REGION Network 11: Habilita cambiar de CAPA_Elem_2
         OPN   "DB_Receta_Actual";
         SET;
         R     #Habil_2_CAPA;
         L     #Capa_Actual;
         L     #Max_Nro_Capas;
         >=I;
         JC    No2CAPA;
         L     #Adress_Capa;
         L     #Length_Capas;
         +I;
         L     #Offset_Filas_DB;
         +I;
         SLD   3;
         L     #Offset_Elementos_DB_bit;
         +I;
         L     #Length_Elementos_DB_bit;
         +I;
         LAR2;
         O     DBX [AR2, P#0.0];
         O     DBX [ AR2 , P#2.0 ];
         =     #Habil_2_CAPA;
   No2CAPA:NOP   0;
END_REGION

REGION Network 12: #Elemento_Actual
         OPN   "DB_Receta_Actual";

         A     DBX [ AR1 , P#4.0 ];
         =     #Elemento_Actual;

         A     #Elemento_Actual;
         JCN   NoActual;
         TAR1  AR2;
END_REGION

REGION Network 13: NUM = 1
         SET;
   // R DBX [ AR1 , P#4.0 ]
         A     #Habil_1_IZQ;
         JCN   No_1_IZQ;

         TAR1  AR2;
         L     1;
         +AR2;
   //S DBX [ AR2 , P#4.0 ]
         JU    Fin;

   No_1_IZQ:A     #Habil_1_ABA;
         JCN   No_ABA;
         L     #Adress_Filas_DB_bit;
         SRD   3;
         L     #Length_Filas_DB;
         +I;
         SLD   3;
         L     #Offset_Elementos_DB_bit;
         +I;
         LAR2;
         SET;
   //S DBX [ AR2 , P#4.0 ]
         JU    Fin;

   No_ABA:A     #Habil_1_CAPA;
         JCN   No_CAPA;
         L     #Adress_Capa;
         L     #Length_Capas;
         +I;
         L     #Offset_Filas_DB;
         +I;
         SLD   3;
         L     #Offset_Elementos_DB_bit;
         +I;
         LAR2;
   //S DBX [ AR2 , P#4.0 ]
         L     #Capa_Actual;
         L     1;
         +I;
         T     #Capa_Actual;
         JU    Fin;

   No_CAPA:NOP   0;
         L     #Offset_Capas;
         L     #Offset_Filas_DB;
         +I;
         SLD   3;
         L     #Offset_Elementos_DB_bit;
         +I;
         LAR2;
   //S DBX [ AR2 , P#4.0 ]
         L     1;
         T     #Capa_Actual;
         L     #Nro_Pallet;
         L     1;
         +I;
         T     #Nro_Pallet;
         JU    Fin;
END_REGION

REGION Network 14: No elemento actual
   NoNUM:JU    Fin;
   NoActual:NOP   0;
END_REGION

REGION Network 15: Bucle Elementos
         L     #Índice_Elementos;
         L     1;
         +I;
         T     #Índice_Elementos;
         L     #Max_Nro_Elementos;
         <=I;
         JC    New_Ele;
END_REGION

REGION Network 16: Bucle Filas
         L     1;
         T     #Índice_Elementos;
         L     #Índice_Filas;
         L     1;
         +I;
         T     #Índice_Filas;
         L     #Max_Nro_Filas;
         <=I;
         JC    New_Fil;
END_REGION

REGION Network 17: #Error
         SET;
         S     #Error;
END_REGION

REGION Network 18: Fin de Bloque
   Fin:  SET;
         R     #Error;
         OPN   "DB_Receta_Actual";
         AN    DBX [ AR2 , P#0.0 ];
         AN    DBX [ AR2 , P#2.0 ];
         JCN   NO_0;
         L     0;
         JU    Transferir;
   NO_0: A     DBX [ AR2 , P#0.0 ];
         AN    DBX [ AR2 , P#2.0 ];
         JCN   NO_1;
         L     1;
         JU    Transferir;
   NO_1: AN    DBX [ AR2 , P#0.0 ];
         A     DBX [ AR2 , P#2.0 ];
         JCN   NO_2;
         L     2;
         JU    Transferir;
   NO_2: L     3;
   Transferir:T     "Proceso Dosificador".Elemento_Proximo;
   // 0 = Invisible
   // 1 = V
   // 2 = H
   // 3 = HH
END_REGION
END_FUNCTION

FUNCTION "FC_Animación" : Void   // FC3, STL
{ S7_Optimized_Access := 'FALSE' }
VERSION : 0.1
BEGIN

REGION Network 1
         O     "Cambio_Elemento";
         O     "flanco"."nHMI.Pls_Inc_Capa";
         O     "flanco"."nHMI.Pls_Dec_Capa";
         O     "flanco"."pHMI.Pls_Inc_Capa_Editando";
         O     "flanco"."pHMI.Pls_Dec_Capa_Editando";

         =     #Cambio_Elemento;
END_REGION

REGION Network 2: Inicializa fila y elemento
         A     "CicIni";
         JCN   L001;
         L     1;
         T     "DB_Animación".Elemento_SEL;
         T     "DB_Animación".Fila_SEL;
         L     "Puntero".Offset_Filas_HMI;
         L     "Puntero".Offset_Elementos_HMI;
         +I;
         SLD   3;
         LAR1;
         OPN   "DB_Animación";
         L     3;
         T     DBB [ AR1 , P#0.0 ];
         S     #Cambio_Elemento;
   L001: NOP   0;

         L     "DB_Animación".Fila_SEL;
         L     "DB_Animación".Elemento_SEL;
   // OFFSET_Y "0" en la primer fila
         L     "Puntero".Offset_Filas_HMI;
         OPN   "DB_Animación";
         SLD   3;
         LAR1;
         L     0;
         T     DBW [ AR1 , P#0.0 ];


   // OFFSET_X "0" en el primer elemento de la primer fila
         L     "Puntero".Offset_Filas_HMI;
         L     "Puntero".Offset_Elementos_HMI;
         +I;
         OPN   "DB_Animación";
         SLD   3;
         LAR1;
         L     0;
         T     DBW [ AR1 , P#2.0 ];

   //Edita recetas
         L     "HMI".Imagen_Actual;
         L     21;
         ==I;
         JC    ED;
         TAK;
         L     22;
         ==I;
         JCN   NoED;
   ED:   S     "Editando_Recetas";
         JU    END;
   NoED: R     "Editando_Recetas";
         S     #Cambio_Elemento;
   END:  NOP   0;
END_REGION

REGION Network 3: Rotación de elemento de Muestra
         L     4;
         L     "DB_Animación".Figura_SEL;
         >I;
         JC    B001;
         L     1;
         T     "DB_Animación".Figura_SEL;
   B001: NOP   0;
         L     "DB_Animación".Figura_SEL;
         T     #Muestra;
END_REGION

REGION Network 4: Inicio Bucle: Recorre elementos HMI
         L     1;
         T     #Índice_Fila;
         T     #Índice_Elemento;

   X001: L     #Índice_Fila;
         L     1;
         -I;
         L     "Puntero".Length_Filas_HMI;
         *I;
         L     "Puntero".Offset_Filas_HMI;
         +I;
         T     #Adress_Fila;
   //Inicio: Nueva fila resetea elementos verticales de la fila
   //        anterior
         R     #No_H;
   //Fin

   X002: L     #Índice_Elemento;
         L     1;
         -I;
         L     "Puntero".Length_Elementos_HMI;
         *I;
         L     "Puntero".Offset_Elementos_HMI;
         +I;
         L     #Adress_Fila;
         +I;
         SLD   3;
         LAR1;

   //Carga en AR2 la dirección del próximo elemento
         SRD   3;
         L     "Puntero".Length_Elementos_HMI;
         +I;
         SLD   3;
         LAR2;







   //   SPA   label
END_REGION

REGION Network 5
   ///////////////////////////////////////////////////////////////
   //                                                           //
   //    INICIO DE BUCLE: A continuación de realizan las        //
   //    tareas para cada elemento, AR1 tiene la dirección      //
   //    del elemento a tratar y AR2 tiene la dirección         //
   //    del siguiente elemento de la fila (ver si existe).     //
   //                                                           //
   ///////////////////////////////////////////////////////////////
   //      SET
   //      S     #Cambio_Elemento


   //Inicio: Se fija en qué dirección se puede mover la selección
   //        de elementos
         OPN   "DB_Animación";
         L     DBB [ AR1,P#1.0];
         L     "Constante".Elemento_SELECCIONADO;
         ==I;
         JCN   NADA;
         TAR2  #Mem_AR2;

   //Habilitar ir hacia la derecha
         L     #Índice_Elemento;
         L     1;
         >I;
         JCN   NoDe;
         CAR;
         LAR1  AR2;
         L     "Puntero".Length_Elementos_HMI;
         SLD   3;
         NEGD;
         +AR2;
         OPN   "DB_Animación";
         L     DBB [ AR2 , P#0.0 ];
         L     0;
         >I;
         =     #Habil_DER;
         JU    SiDe;
   NoDe: R     #Habil_DER;
   SiDe: NOP   0;

   //Habilitar ir hacia la izquierda
         L     #Índice_Elemento;
         L     "Puntero".Max_Nro_Elementos;
         <I;
         JCN   NoIz;
         CAR;
         LAR1  AR2;
         L     "Puntero".Length_Elementos_HMI;
         SLD   3;
         +AR2;
         OPN   "DB_Animación";
         L     DBB [ AR2 , P#0.0 ];
         L     0;
         >I;
         =     #Habil_IZQ;
         JU    SiIz;
   NoIz: R     #Habil_IZQ;
   SiIz: NOP   0;



   //Habilitar ir hacia arriba
         L     #Índice_Fila;
         L     1;
         >I;
         JCN   NoSu;
         CAR;
         LAR1  AR2;
         L     "Puntero".Length_Filas_HMI;
         SLD   3;
         NEGD;
         +AR2;
         OPN   "DB_Animación";
         L     DBB [ AR2 , P#0.0 ];
         L     0;
         >I;
         =     #Habil_SUBIR;
         JU    SiSu;
   NoSu: R     #Habil_SUBIR;
   SiSu: NOP   0;

   //Habilitar ir hacia abajo
         L     #Índice_Fila;
         L     "Puntero".Max_Nro_Filas;
         <I;
         JCN   NoBa;
         CAR;
         LAR1  AR2;
         L     "Puntero".Length_Filas_HMI;
         SLD   3;
         +AR2;
         OPN   "DB_Animación";
         L     DBB [ AR2 , P#0.0 ];
         L     0;
         >I;
         =     #Habil_BAJAR;
         JU    SiBa;
   NoBa: R     #Habil_BAJAR;
   SiBa: NOP   0;
END_REGION

REGION Network 6: Recorre elementos HMI
   //Inicio: Si no está en modo de edición de recetas, fuerza el cambio de
   //        de selección si hubo un "Elemento_CARGADO".
         A     "Editando_Recetas";
         JC    edit;
         A     "Elemento_CARGADO";
         A     #Habil_IZQ;
         JCN   c1;
         L     "DB_Animación".Elemento_SEL;
         INC   1;
         T     "DB_Animación".Elemento_SEL;
         S     #Cambio_Elemento;
         R     "Elemento_CARGADO";
         JU    edit;

   //Se fija si puede haber una fila más abajo
   c1:   L     #Índice_Fila;
         L     "Puntero".Max_Nro_Filas;
         <I;
         JCN   edit;
   //Se fija si el primer elemento de la fila inferior existe
         L     #Adress_Fila;
         L     "Puntero".Length_Filas_HMI;
         +I;
         L     "Puntero".Offset_Elementos_HMI;
         +I;
         SLD   3;
         LAR2;
         OPN   "DB_Animación";
         L     DBB [AR2,P#0.0];
         L     0;
         <>I;
         A     "Elemento_CARGADO";
         JCN   c22;
         L     "DB_Animación".Fila_SEL;
         INC   1;
         T     "DB_Animación".Fila_SEL;
         L     1;
         T     "DB_Animación".Elemento_SEL;
         S     #Cambio_Elemento;
         R     "Elemento_CARGADO";
         JU    edit;
   c22:  A     "Elemento_CARGADO";
         A     "CICLO_Hab";
         JCN   edit;
         =     "Nueva_CAPA";
         L     1;
         T     "DB_Animación".Elemento_SEL;
         T     "DB_Animación".Fila_SEL;
         S     #Cambio_Elemento;
         R     "Elemento_CARGADO";
   edit: NOP   0;
   //Fin

















   //Inicio: Si no está en modo de edición de recetas, fuerza el cambio de
   //        selección si hubo un "Elemento_DESCARGADO".

         O     "Editando_Recetas";
         ON    "Elemento_DESCARGADO";
         JC    Final;
         A     #Habil_DER;
         JCN   FILA;
         L     "DB_Animación".Elemento_SEL;
         DEC   1;
         T     "DB_Animación".Elemento_SEL;
         S     #Cambio_Elemento;
         R     "Elemento_DESCARGADO";
         JU    Final;

   //Se fija si puede haber una fila más arriba
   FILA: L     #Adress_Fila;
         L     1;
         >I;
         JCN   Final;
   //Elije el último elemento que exista de la fila superior
         L     #Adress_Fila;
         L     "Puntero".Length_Filas_HMI;
         -I;
         L     "Puntero".Offset_Elementos_HMI;
         +I;
         L     "Puntero".Length_Elementos_HMI;
         -I;
         T     #Temp;
   NO_Cero:L     #Temp;
         L     "Puntero".Length_Elementos_HMI;
         +I;
         T     #Temp;
         SLD   3;
         LAR2;
         OPN   "DB_Animación";
         L     DBB [AR2,P#0.0];
         L     0;
         ==I;
         JCN   NO_Cero;
         L     #Temp;
         L     "Puntero".Offset_Elementos_HMI;
         -I;
         L     #Adress_Fila;
         -I;
         L     "Puntero".Length_Filas_HMI;
         +I;

         L     "Puntero".Length_Elementos_HMI;
         /I;
         T     "DB_Animación".Elemento_SEL;
         L     "DB_Animación".Fila_SEL;
         DEC   1;
         T     "DB_Animación".Fila_SEL;
         S     #Cambio_Elemento;
   Final:R     "Elemento_DESCARGADO";

   //Fin













   //
         LAR2  #Mem_AR2;
   //



   //Se fija si hay que mover el elemento seleccionado hacia
   //la derecha
         A     "flanco".piPul_MultiAde;
         A     #Habil_DER;
         A     "Editando_Recetas";
         JCN   A001;
   //   SET

         S     #Cambio_Elemento;
         L     "DB_Animación".Elemento_SEL;
         DEC   1;
         T     "DB_Animación".Elemento_SEL;
         JC    A004;
   //Se fija si hay que mover el elemento seleccionado hacia
   //la izquierda
   A001: A     "flanco".piPul_MultiAtr;
         A     #Habil_IZQ;
         A     "Editando_Recetas";
         JCN   A002;
   //   SET

         S     #Cambio_Elemento;
         L     "DB_Animación".Elemento_SEL;
         INC   1;
         T     "DB_Animación".Elemento_SEL;
         JC    A004;
   //Se fija si hay que mover el elemento seleccionado hacia
   //arriba
   A002: A     "flanco".piPul_MultiArr;
         A     #Habil_SUBIR;
         A     "Editando_Recetas";
         JCN   A003;
   //    SET

         S     #Cambio_Elemento;
         L     "DB_Animación".Fila_SEL;
         DEC   1;
         T     "DB_Animación".Fila_SEL;
         JC    A004;
   //Se fija si hay que mover el elemento seleccionado hacia
   //abajo
   A003: A     "flanco".piPul_MultiAba;
         A     #Habil_BAJAR;
         A     "Editando_Recetas";
         JCN   A004;
   //    SET

         S     #Cambio_Elemento;
         L     "DB_Animación".Fila_SEL;
         INC   1;
         T     "DB_Animación".Fila_SEL;
   //Se fija si hubo un cambio en el elemento seleccionado
   A004: NOP   0;
   //   O     "Elemento_CARGADO"
   //   O     "Elemento_DESCARGADO"
   //   =     #Cambio_Elemento
   //
   //    R     "Elemento_CARGADO"
   //    R     "Elemento_DESCARGADO"
   NADA: NOP   0;
   //      SET
   //      S     #Cambio_Elemento
   //Fin
END_REGION

REGION Network 7: "S_PriElemCapa"
         OPN   "DB_Animación";
         L     DBB [ AR1,P#1.0];
         L     "Constante".Elemento_SELECCIONADO;
         ==I;
         JCN   PriElem;
         L     #Índice_Elemento;
         L     1;
         ==I;
         JCN   NoPriElem;
         L     #Índice_Fila;
         ==I;
         S     "S_PriElemCapa";
         JU    PriElem;
   NoPriElem:R     "S_PriElemCapa";
   PriElem:NOP   0;
END_REGION

REGION Network 8: Recorre elementos HMI: Kill_Elemento
   //Inicio: Hacer que el elemento seleccionado tenga figura "0",
   //        es decir, que desaparezca.
         OPN   "DB_Animación";
         L     DBB [ AR1,P#1.0];
         L     "Constante".Elemento_SELECCIONADO;
         ==I;
         JCN   J001;
         A     "flanco"."pHMI.Pls_Kill_Elem";
         JCN   J001;
         L     #Índice_Elemento;
         L     1;
         ==I;
         JCN   J002;
         L     #Índice_Fila;
         ==I;
         JC    J001;

   J002: L     0;
         OPN   "DB_Animación";
         T     DBB [ AR1,P#0.0];
   J001: NOP   0;
   //Fin

   //Inicio: Hacer que si el elemento seleccionado tiene figura "0",
   //        o sea, no existe, la selección cambie al elemento
   //        anterior de la fila o al elemento 1 de la fila anterior.
         OPN   "DB_Animación";
         L     DBB [ AR1 , P#1.0 ];
         L     "Constante".Elemento_SELECCIONADO;
         ==I;
         JCN   J003;
         OPN   "DB_Animación";
         L     DBB [ AR1 , P#0.0 ];
         L     0;
         ==I;
         JCN   J003;
         L     #Índice_Elemento;
         L     1;
         >I;
         JCN   J004;
         L     "DB_Animación".Elemento_SEL;
         DEC   1;
         T     "DB_Animación".Elemento_SEL;
         S     #Cambio_Elemento;
         JU    J003;
   J004: L     "DB_Animación".Fila_SEL;
         DEC   1;
         T     "DB_Animación".Fila_SEL;
         S     #Cambio_Elemento;
   J003: NOP   0;
   //Fin
END_REGION

REGION Network 9: Recorre elementos HMI: New_Elemento
   //Inicio: Si el elemento tiene figura "0" (invisible) y el elemento
   //        anterior de la fila tiene figura <> "0", copia la figura
   //        del elemento anterior. Esto si el elemento actual no es
   //        el primero de la fila.
         OPN   "DB_Animación";
         L     #Índice_Fila;
         L     "DB_Animación".Fila_SEL;
         ==I;
         JCN   D001;
         OPN   "DB_Animación";
         L     DBB [ AR1 , P#0.0 ];
         L     0;
         ==I;
         JCN   D001;
         L     #Índice_Elemento;
         L     1;
         >I;
         A     "flanco"."pHMI.Pls_New_Elem";
         JCN   D001;
         TAR2  #Mem_AR2;
         CAR;
         LAR1  AR2;
         L     "Puntero".Length_Elementos_HMI;
         SLD   3;
         NEGD;
         +AR2;
         OPN   "DB_Animación";
         L     0;
         L     DBB[AR2,P#0.0];
         <I;
         JCN   D001;
         T     DBB [ AR1 , P#0.0 ];
         R     "flanco"."pHMI.Pls_New_Elem";
         LAR2  #Mem_AR2;
   D001: OPN   "DB_Animación";
   //Fin
END_REGION

REGION Network 10: Recorre elementos HMI: New_Fila
   //Inicio: Si el elemento tiene figura "0" (invisible), es el primer
   //        elemento de la fila, y el primer elemento de la fila anterior
   //        tiene figura <> "0", copia la figura de aquel elemento.
         OPN   "DB_Animación";
         L     #Índice_Fila;
         L     "Puntero".Max_Nro_Filas;
         <=I;
         JCN   E001;
         OPN   "DB_Animación";
         L     DBB [ AR1 , P#0.0 ];
         L     0;
         ==I;
         JCN   E001;
         L     #Índice_Elemento;
         L     1;
         ==I;
         A     "flanco"."pHMI.Pls_New_Fila";
         JCN   E001;
         TAR2  #Mem_AR2;
         CAR;
         LAR1  AR2;
         L     "Puntero".Length_Filas_HMI;
         SLD   3;
         NEGD;
         +AR2;
         OPN   "DB_Animación";
         L     0;
         L     DBB[AR2,P#0.0];
         <I;
         JCN   E001;
         T     DBB [ AR1 , P#0.0 ];
         R     "flanco"."pHMI.Pls_New_Fila";
         LAR2  #Mem_AR2;
   E001: OPN   "DB_Animación";




   //Fin
END_REGION

REGION Network 11: Recorre elementos HMI: Maca elemento seleccionado
   //Inicio: Marca elemento como seleccionado y
   //        desmarca todos los otros
         OPN   "DB_Animación";
         L     #Índice_Fila;
         L     "DB_Animación".Fila_SEL;
         <=I;
         JCN   X013;
         >=I;
         JCN   x014;

         L     #Índice_Elemento;
         L     "DB_Animación".Elemento_SEL;
         <=I;
         JCN   X013;
         >=I;
         JCN   x014;
         L     "Constante".Elemento_SELECCIONADO;
         OPN   "DB_Animación";
         T     DBB [ AR1 , P#1.0];

   //Inicio: Si hubo cambio de selección copia la figura
   //        del elemento seleccionado.
         O     #Cambio_Elemento;
         O     "flanco".pEditando_Recetas;
   //  O     "flanco"."pHMI.Pls_RD_Receta"
   //
         OPN   "DB_Animación";
         JCN   X006;
         L     DBB [ AR1 , P#0.0 ];
         T     #Muestra;
         SET;
         R     #Cambio_Elemento;
   X006: L     #Muestra;
         T     DBB [ AR1 , P#0.0 ];
   //Fin
         JU    X005;
   X013: A     "Editando_Recetas";
         JC    x014;
         L     "Constante".Elemento_AUSENTE;
         JU    X004;
   x014: L     "Constante".Elemento_PRESENTE;  //Estado de elementos no seleccionado

   X004: OPN   "DB_Animación";
         T     DBB [ AR1 , P#1.0 ];
   X005: NOP   0;
   //Fin
END_REGION

REGION Network 12: Recorre elementos HMI: Borra elementos

   //Inicio: Si es "0" (invisible) la figura del elemento 1 de la fila,
   //        pone a "0" el elemento 1 de la fila siguiente (si la hay)
         L     #Índice_Fila;
         L     "Puntero".Max_Nro_Filas;
         OPN   "DB_Animación";
         <I;
         JCN   C001;
         L     #Índice_Elemento;
         L     1;
         ==I;
         JCN   C001;
         L     DBB [ AR1 , P#0.0 ];
         L     0;
         ==I;
         JCN   C001;
         TAR2  #Mem_AR2;
         CAR;
         LAR1  AR2;
         L     "Puntero".Length_Filas_HMI;
         OPN   "DB_Animación";
         SLD   3;
         +AR2;
         TAK;
         T     DBB [ AR2 , P#0.0 ];
         LAR2  #Mem_AR2;
   C001: NOP   0;
   //Fin

   //Inicio: Si la figura del elemento actual es "0" (invisible)
   //        pone a "0" la figura del elemento siguiente
   //        en la misma fila (Si lo hay)
         L     #Índice_Elemento;
         L     "Puntero".Max_Nro_Elementos;
         >=I;
         JC    X012;
         OPN   "DB_Animación";
         L     DBB [ AR1 , P#0.0 ];
         L     0;
         <>I;
         JC    X012;
         T     DBB [ AR2 , P#0.0 ];
   X012: NOP   0;
   //Fin
END_REGION

REGION Network 13: Recorre elementos HMI
   //Forzar la figura de los elementos para probar
         OPN   "DB_Animación";
   //      L     3
   //      T DBB [ AR1 , P#0.0 ]
   //Forzar lOffset de los elementos para probar
         OPN   "DB_Animación";
   //     L     0
   //     T DBW [ AR1 , P#2.0 ]



   //Inicio: Revisa si hay algún elemento que no sea horizontal (Figura 2)
   //        en la fila actual, para ajustar Offset_Y
         OPN   "DB_Animación";
         L     DBB [ AR1 , P#0.0 ];
         L     2;
         ==I;
         JC    X009;
         TAK;
         L     0;
         ==I;
         JC    X009;
         S     #No_H;
   X009: NOP   0;
   //Fin


   //Inicio: Offset elemento siguiente en función del Offset y la
   //        figura del elemento actual
         L     #Índice_Elemento;
         L     "Puntero".Max_Nro_Elementos;
         >=I;
         JC    X008;
         OPN   "DB_Animación";
         L     DBB [ AR1 , P#0.0 ];
         L     1;
         <=I;
         JC    X007;
         L     DBW [ AR1 , P#2.0 ];
         L     "Constante".HMI_Pixel_Offset_X;
         +I;
         OPN   "DB_Animación";
         T     DBW [ AR2 , P#2.0 ];
         JU    X008;
   X007: L     DBW [ AR1 , P#2.0 ];
         T     DBW [ AR2 , P#2.0 ];
   X008: NOP   0;
   //Fin

   //Inicio: Si no es la primer fila, ajusta Offset_Y dependiendo
   //        de si tiene sólo elementos "H" (Figura 2) o no.
         TAR1  #Mem_AR1;
         TAR2  #Mem_AR2;
         L     #Adress_Fila;
         SLD   3;
         LAR1;
         L     #Índice_Fila;
         L     1;
         <=I;
         JC    X011;
   //Carga en AR2 la dirección de la fila anterior
         L     #Adress_Fila;
         L     "Puntero".Length_Filas_HMI;
         -I;
         SLD   3;
         LAR2;

         OPN   "DB_Animación";
         AN    #No_H;
         JC    X010;
         L     DBW [ AR2 , P#0.0 ];
         L     "Constante".HMI_Pixel_Offset_Y;
         +I;
         OPN   "DB_Animación";
         T     DBW [ AR1 , P#0.0 ];
         JU    X011;
   X010: L     DBW [ AR2 , P#0.0 ];
         T     DBW [ AR1 , P#0.0 ];
   X011: NOP   0;
         LAR1  #Mem_AR1;
         LAR2  #Mem_AR2;
   //Fin
END_REGION

REGION Network 14: Señales2
   //
         AN    #Habil_IZQ;
         =     "S_ÚltElemFila";

   //
         TAR1  #Mem_AR1;
         TAR2  #Mem_AR2;

         OPN   "DB_Animación";
         L     DBB [ AR1,P#1.0];
         L     "Constante".Elemento_SELECCIONADO;
         ==I;
         JCN   NoUltFil2;

         L     #Índice_Fila;
         L     "Puntero".Max_Nro_Filas;
         <I;
         JCN   Ult_Fil;
   //Carga en AR2 la dirección de la fila posterior
         L     #Adress_Fila;
         L     "Puntero".Length_Filas_HMI;
         +I;
         SLD   3;
         LAR2;
   //
   //Calcula en AR2 la dirección del primer elemento
         L     "Puntero".Offset_Elementos_HMI;
         SLD   3;
         +AR2;
   //
   Ult_Fil:NOP   0;

         O(;
         L     #Índice_Fila;
         L     "Puntero".Max_Nro_Filas;
         ==I;
         );
         O(;
         A(;
         L     #Índice_Fila;
         L     "Puntero".Max_Nro_Filas;
         <I;
         );
         A(;
         OPN   "DB_Animación";
         L     DBB [ AR2 , P#0.0 ];
         L     "Constante".Elemento_AUSENTE;
         ==I;
         );
         );
         =     "S_ÚltFilCapa";
   NoUltFil2:NOP   0;

         LAR1  #Mem_AR1;
         LAR2  #Mem_AR2;

   // NO anduvo
   //     U     "S_ÚltFilCapa"
   //      U     "iSnsEmpj_Ade_Par"
   //     U     "iSnsEmpj_Arriba"
   //     R     "S_ÚltFilCapa"
END_REGION

REGION Network 15
   label:NOP   0;
   ///////////////////////////////////////////////////////////////
   //                                                           //
   //    FIN DE BUCLE:                                          //
   //                                                           //
   ///////////////////////////////////////////////////////////////
END_REGION

REGION Network 16: Fin Bucle: Recorre elementos HMI
         L     #Índice_Elemento;
         L     1;
         +I;
         T     #Índice_Elemento;
         L     "Puntero".Max_Nro_Elementos;
         <=I;
         JC    X002;
         L     1;
         T     #Índice_Elemento;
         L     #Índice_Fila;
         L     1;
         +I;
         T     #Índice_Fila;
         L     "Puntero".Max_Nro_Filas;
         <=I;
         JC    X001;
END_REGION

REGION Network 17
         L     #Muestra;
         T     "DB_Animación".Figura_SEL;
   //
         A     #Cambio_Elemento;
         =     "Cambio_Elemento";
   //
   //   R     "HMI".Pls_RD_Receta
END_REGION
END_FUNCTION

FUNCTION "CAPA Receta_Animación_Receta" : Void   // FC6, STL
{ S7_Optimized_Access := 'FALSE' }
VERSION : 0.1
BEGIN

REGION Network 1
         CLR;
         =     #Reset_RD_Receta;
   //Resetear Nro_Receta_Edición y Capa_Actual_Edición
         A     "flanco".pEditando_Recetas;
         JCN   Edita1;
         L     1;
   // T     "DB_Animación".Nro_Receta_Edición
         T     "DB_Animación".Capa_Actual_Edición;
   Edita1:NOP   0;
   //
         O     "xpEditar_Recetas";
         O     "flanco"."nHMI.Pls_RD_Receta";
         JCN   Salir;
END_REGION

REGION Network 2: Modifica RECETA

         JC    NO2R;
   //Incrementar Receta_EDITANDO
         L     "DB_Animación".Nro_Receta_Edición;
         L     10;
         <I;
         JCN   RMax;
         A     "flanco"."nHMI.Pls_Inc_Receta";
         JCN   NO1R;
         L     "DB_Animación".Nro_Receta_Edición;
         L     1;
         +I;
         T     "DB_Animación".Nro_Receta_Edición;
         JU    NO1R;
   RMax: L     10;
         T     "DB_Animación".Nro_Receta_Edición;
   NO1R: NOP   0;
   //Decrementar Receta_EDITANDO
         L     "DB_Animación".Nro_Receta_Edición;
         L     1;
         >I;
         JCN   RMin;
         A     "flanco"."nHMI.Pls_Dec_Receta";
         JCN   NO2R;
         L     "DB_Animación".Nro_Receta_Edición;
         L     1;
         -I;
         T     "DB_Animación".Nro_Receta_Edición;
         JU    NO2R;
   RMin: L     1;
         T     "DB_Animación".Nro_Receta_Edición;
   NO2R: NOP   0;
END_REGION

REGION Network 3: Modifica CAPA

         JCN   NO2C;
   //Incrementar Capa_EDITANDO
         L     "DB_Animación".Capa_Actual_Edición;
         L     10;  //  L     "Proceso Dosificador".CapasDistinReceta
         <I;
         JCN   CMax;
         A     "flanco"."pHMI.Pls_Inc_Capa_Editando";
         JCN   NO1C;
         L     "DB_Animación".Capa_Actual_Edición;
         L     1;
         +I;
         T     "DB_Animación".Capa_Actual_Edición;
         JU    NO1C;
   CMax: NOP   0;  // L     "Proceso Dosificador".CapasDistinReceta
         T     "DB_Animación".Capa_Actual_Edición;
   NO1C: NOP   0;
   //Decrementar Capa_EDITANDO
         L     "DB_Animación".Capa_Actual_Edición;
         L     1;
         >I;
         JCN   CMin;
         A     "flanco"."pHMI.Pls_Dec_Capa_Editando";
         JCN   NO2C;
         L     "DB_Animación".Capa_Actual_Edición;
         L     1;
         -I;
         T     "DB_Animación".Capa_Actual_Edición;
         JU    NO2C;
   CMin: L     1;
         T     "DB_Animación".Capa_Actual_Edición;
   NO2C: NOP   0;
END_REGION

REGION Network 4: Constantes
         L     "DB_Animación".Nro_Receta_Edición;
         T     #Receta_Actual;
         L     "Puntero".Length_Recetas;
   //    L     312
         T     #Length_Recetas;
         L     "Puntero".Offset_Recetas;
   //    L     0
         T     #Offset_Recetas;
         L     "DB_Animación".Capa_Actual_Edición;
         T     #Capa_Actual;
         L     "Puntero".Length_Capas_Receta;
   //    L     26
         T     #Length_Capas;
         L     "Puntero".Offset_Capas_Receta;
   //    L     52
         T     #Offset_Capas;
         L     "Puntero".Length_Filas_CapaReceta;
   //    L     4
         T     #Length_Filas_DB;
         L     "Puntero".Offset_Filas_CapaReceta;
   //    L     0
         T     #Offset_Filas_DB;
         L     1;
         T     #Length_Elementos_DB_bit;
         L     0;
         T     #Offset_Elementos_DB_bit;

         L     1;
         T     #Índice_Filas;
         T     #Índice_Elementos;

         SET;
         R     #f_Selec;

         L     "Puntero".Length_Filas_HMI;
         T     #Length_Filas_DI;
         L     "Puntero".Offset_Filas_HMI;
         T     #Offset_Filas_DI;
         L     "Puntero".Length_Elementos_HMI;
         T     #Length_Elementos_DI;
         L     "Puntero".Offset_Elementos_HMI;
         T     #Offset_Elementos_DI;

         L     "Constante".Elemento_PRESENTE;
         T     #Elemento_Cargado;
         L     "Constante".Elemento_SELECCIONADO;
         T     #Elemento_Siguiente;
         L     "Constante".Elemento_AUSENTE;
         T     #Elemento_Ausente;

         L     "Puntero".Max_Nro_Elementos;
         T     #Max_Nro_Elementos;
         L     "Puntero".Max_Nro_Filas;
         T     #Max_Nro_Filas;
END_REGION

REGION Network 5: #Adress_Receta
         L     #Receta_Actual;
         L     1;
         -I;
         L     #Length_Recetas;
         *I;
         L     #Offset_Recetas;
         +I;
         T     #Adress_Receta;
END_REGION

REGION Network 6: Adress_Capa
         L     #Capa_Actual;
         L     1;
         -I;
         L     #Length_Capas;
         *I;
         L     #Offset_Capas;
         +I;
         L     #Adress_Receta;
         +I;
         T     #Adress_Capa;
END_REGION

REGION Network 7
         TAR1  #Mem_AR1;  // Memorizar AR1
         TAR2  #Mem_AR2;  // Memorizar AR2
         T     #Mem_Accu1;  // Memorizar Accu1
         TAK;
         T     #Mem_Accu2;  // Memorizar Accu2
   //################################################

         L     #Adress_Capa;
         L     24;  // Offset Usar Pistón
         +I;
         SLD   3;
         LAR1;

   // Si no hubo cambio de capa, del gráfico a la receta
         AN    "flanco"."pHMI.Pls_Inc_Capa_Editando";
         AN    "flanco"."pHMI.Pls_Dec_Capa_Editando";
         AN    "HMI".Pls_RD_Receta;
         JCN   NoEditar;

         A     "DB_Animación".Usar_Pistón;
         OPN   "DB_RECETAS";
         =     DBX [ AR1 ,P#0.0];
   NoEditar:NOP   0;

   // De la receta al gráfico
         OPN   "DB_RECETAS";
         A     DBX [ AR1 , P#0.0 ];
         =     "DB_Animación".Usar_Pistón;

   //################################################
         L     #Mem_Accu2;  // Recuperar Accu2
         L     #Mem_Accu1;  // Recuperar Accu1
         LAR1  #Mem_AR1;  // Recuperar AR1
         LAR2  #Mem_AR2;  // Recuperar AR2
END_REGION

REGION Network 8: Adress_Filas_DB
   New_Fil:NOP   0;
         L     #Índice_Filas;
         L     1;
         -I;
         L     #Length_Filas_DB;
         *I;
         L     #Offset_Filas_DB;
         +I;
         L     #Adress_Capa;
         +I;
         SLD   3;
         T     #Adress_Filas_DB_bit;
END_REGION

REGION Network 9: Adress_Filas_DI
         L     #Índice_Filas;
         L     1;
         -I;
         L     #Length_Filas_DI;
         *I;
         L     #Offset_Filas_DI;
         +I;
         T     #Adress_Filas_DI;
END_REGION

REGION Network 10: Adress_Elementos_DB
   New_Ele:NOP   0;
         L     #Índice_Elementos;
         L     1;
         -I;
         L     #Length_Elementos_DB_bit;
         *I;
         L     #Offset_Elementos_DB_bit;
         +I;
         L     #Adress_Filas_DB_bit;
         +I;
         T     #Adress_Elementos_DB_bit;
END_REGION

REGION Network 11: Adress_Elementos_DI
         L     #Índice_Elementos;
         L     1;
         -I;
         L     #Length_Elementos_DI;
         *I;
         L     #Offset_Elementos_DI;
         +I;
         L     #Adress_Filas_DI;
         +I;
         T     #Adress_Elementos_DI;
END_REGION

REGION Network 12: AR1 y AR2
         L     #Adress_Elementos_DB_bit;
         LAR1;
         L     #Adress_Elementos_DI;
         SLD   3;
         LAR2;
END_REGION

REGION Network 13: Transferencia de Figuras
   // Si no hay cambio de capa, transfiere del gráfico a la receta
         L     "HMI".Imagen_Actual;
         L     22;
         ==I;
         L     S5T#30S;
         SD    "Tag_1";
         A     "Tag_1";
         AN    "flanco"."pHMI.Pls_Inc_Capa_Editando";
         AN    "flanco"."pHMI.Pls_Dec_Capa_Editando";
         AN    "HMI".Pls_RD_Receta;

         JCN   Fin;
   //SPA   Fin

         OPN   "DB_RECETAS";
         OPNDI "DB_Animación";
   // 0 = Invisible
   // 1 = V
   // 2 = H
   // 3 = HH
         L     DIB [ AR2 , P#0.0 ];
         L     0;
         ==I;
         JCN   NO_00;
         R     DBX[AR1,P#0.0];
         R     DBX [ AR1 , P#2.0 ];
         JU    Fin;
   NO_00:L     DIB [ AR2 , P#0.0 ];
         L     1;
         ==I;
         JCN   NO_10;
         S     DBX [ AR1 , P#0.0 ];
         R     DBX [ AR1 , P#2.0 ];
         JU    Fin;
   NO_10:L     DIB [ AR2 , P#0.0 ];
         L     2;
         ==I;
         JCN   NO_20;
         R     DBX[AR1,P#0.0];
         S     DBX [ AR1 , P#2.0 ];
         JU    Fin;
   NO_20:S     DBX [ AR1 , P#0.0 ];
         S     DBX [ AR1 , P#2.0 ];
   Fin:  NOP   0;
END_REGION

REGION Network 14: Transferencia de Figuras
   // Transfiere de la receta al gráfico

         OPN   "DB_RECETAS";
         OPNDI "DB_Animación";
   // 0 = Invisible
   // 1 = V
   // 2 = H
   // 3 = HH

         AN    DBX [ AR1 , P#0.0 ];
         AN    DBX [ AR1 , P#2.0 ];
         JCN   NO_0;
         L     0;
         JU    Transferir;
   NO_0: A     DBX [ AR1 , P#0.0 ];
         AN    DBX [ AR1 , P#2.0 ];
         JCN   NO_1;
         L     1;
         JU    Transferir;
   NO_1: AN    DBX [ AR1 , P#0.0 ];
         A     DBX [ AR1 , P#2.0 ];
         JCN   NO_2;
         L     2;
         JU    Transferir;
   NO_2: L     3;
   Transferir:T     DIB [ AR2 , P#0.0 ];
END_REGION

REGION Network 15: Bucle Elementos
         L     #Índice_Elementos;
         L     1;
         +I;
         T     #Índice_Elementos;
         L     #Max_Nro_Elementos;
         <=I;
         JC    New_Ele;
END_REGION

REGION Network 16: Bucle Filas
         L     1;
         T     #Índice_Elementos;
         L     #Índice_Filas;
         L     1;
         +I;
         T     #Índice_Filas;
         L     #Max_Nro_Filas;
         <=I;
         JC    New_Fil;
END_REGION

REGION Network 17: Fin de Bloque
   Salir:NOP   0;
   // R     "HMI".Pls_RD_Receta
         BEU;
END_REGION
END_FUNCTION

FUNCTION "FC_CARGA_RECETA" : Void   // FC17, STL
TITLE = Carga los datos de la receta seleccionada en Receta Actual y genera las capas correspondientes
{ S7_Optimized_Access := 'FALSE' }
VERSION : 0.1
BEGIN

REGION Network 1: Carga de constantes
   //Carga de constantes
         L     "Puntero".Offset_Recetas;
         T     #Offset_Recetas;
         L     "Puntero".Length_Recetas;
         T     #Length_Recetas;
         L     "Puntero".Offset_Nombre_Receta;
         T     #Offset_Nombre_Receta_DB;
         L     "Puntero".Length_Capas_Receta;
         T     #Length_Capas_DB;
         L     "Puntero".Offset_Capas_Receta;
         T     #Offset_Capas_DB;
         L     "Puntero".Length_Filas_CapaReceta;
         T     #Length_Filas_CapaReceta_DB;
         L     "Puntero".Offset_Filas_CapaReceta;
         T     #Offset_Filas_CapaReceta_DB;
         L     "Puntero".Offset_CapasDist_Receta;
   //    L     51
         T     #Offset_CapasDist_Receta_DB;
         L     "Puntero".Offset_CantCapas_Receta;
   //    L     50
         T     #Offset_CantCapas_Receta_DB;
         L     "Puntero".Offset_Vel_Dosificador;
         T     #Offset_Vel_Dosificador;
         L     "Puntero".Length_Vel_Dosificador;
         T     #Length_Vel_Dosificador;

   //
         L     "Puntero".Length_Nombre_Receta;
   //    L     50
         T     #Length_Nombre_Receta;
   //

         L     52;
         T     #Offset_CantCapas_Receta_DI;
         L     53;
         T     #Offset_CapasDist_Receta_DI;
         L     54;
         T     #Offset_Capas_DI;
         L     6;
         T     #Length_Filas_CapaReceta_DI;
         L     38;
         T     #Length_Capas_DI;
         L     0;
         T     #Offset_Filas_CapaReceta_DI;
   //
         L     "Puntero".Max_Nro_Filas;
         T     #Max_Nro_Filas;
         L     "Puntero".Max_Nro_Elementos;
         T     #Max_Nro_Elementos;
         L     "Puntero".Max_Nro_Capas;
         T     #Max_Nro_Capas;
         L     0;
         T     #índice_Capa_DB;
         T     #Índice_Capa_DI;
         T     #"Nro CapaActual";

         SET;
         R     #Reset_Bit;
         S     #Primer_Elemento;
END_REGION

REGION Network 2: Abrir la receta correspondiente
         L     #"NRO RECETA";
         DEC   1;
         L     #Length_Recetas;
         *I;
         L     #Offset_Recetas;
         +I;
         T     #Adress_Receta;
END_REGION

REGION Network 3: Transferir Número de receta

         L     #"NRO RECETA";
         T     "DB_Receta_Actual".Número;
END_REGION

REGION Network 4: Transferir Nombre de receta

         OPN   "DB_RECETAS";
         OPNDI "DB_Receta_Actual";
         L     #Adress_Receta;
         L     #Offset_Nombre_Receta_DB;
         +I;
         SLD   3;
         LAR1;
         L     2;
         SLD   3;
         LAR2;
         L     0;
         T     #K;
   Bucle:SLD   3;
         OPN   "DB_RECETAS";
         OPNDI "DB_Receta_Actual";
         +AR1;
         +AR2;
         L     DBB [ AR1 , P#0.0 ];
         T     DIB [ AR2 , P#0.0 ];
         L     #K;
         INC   1;
         T     #K;
         L     #Length_Nombre_Receta;
         <I;
         L     1;
         JC    Bucle;
END_REGION

REGION Network 5: Transferir Número de capas por pallet
         OPN   "DB_RECETAS";
         OPNDI "DB_Receta_Actual";
         L     #Adress_Receta;
         L     #Offset_CantCapas_Receta_DB;
         +I;
         SLD   3;
         LAR1;
         L     #Offset_CantCapas_Receta_DI;
         SLD   3;
         LAR2;
         L     DBB [AR1, P#0.0];
         T     DIB [ AR2 , P#0.0 ];
         T     #Nro_Capas;
END_REGION

REGION Network 6: Transferir Número de capas distintas
         OPN   "DB_RECETAS";
         OPNDI "DB_Receta_Actual";
         L     #Adress_Receta;
         L     #Offset_CapasDist_Receta_DB;
         +I;
         SLD   3;
         LAR1;
         L     #Offset_CapasDist_Receta_DI;
         SLD   3;
         LAR2;
         L     DBB [AR1, P#0.0];
         T     DIB [ AR2 , P#0.0 ];
         T     #Nro_CapasDistintas;
END_REGION

REGION Network 7: Completar formato pallet a partir de la receta
   //SPA   m000
         OPN   "DB_RECETAS";
         OPNDI "DB_Receta_Actual";
   Bucle_3:L     #índice_Capa_DB;
         L     #Length_Capas_DB;
         *I;
         L     #Offset_Capas_DB;
         +I;
         L     #Adress_Receta;  // Adress_Receta
         +I;
         T     #Adress_Capa_DB;  // Adress_Capa

         L     #Offset_Filas_CapaReceta_DB;
         +I;
         T     #Adress_Fila_DB;  // Adress_Fila
         SLD   3;
         LAR1;  //Dirección fila
         L     #Índice_Capa_DI;
         L     #Length_Capas_DI;
         *I;
         L     #Offset_Capas_DI;
         +I;
         T     #Adress_Capa_DI;

         L     #Offset_Filas_CapaReceta_DI;
         +I;
         T     #Adress_Fila_DI;
         SLD   3;
         LAR2;  //Dirección fila

         L     0;
         T     #Contador_Filas;
         T     #Contador_Elementos;

   //Transferencia del bit "Usar_Pistón" a la receta actual
   //  SPA   next
         TAR1  #Mem_AR1;  // Memorizar AR1
         TAR2  #Mem_AR2;  // Memorizar AR2
         T     #Mem_Accu1;
         TAK;
         T     #Mem_Accu2;

         L     #Adress_Capa_DB;
         L     24;
         +I;
         SLD   3;
         LAR1;

         L     #Adress_Capa_DI;
         L     36;
         +I;
         SLD   3;
         LAR2;

         OPN   "DB_RECETAS";
         OPNDI "DB_Receta_Actual";
         A     DBX [ AR1 , P#0.0 ];
         =     DIX [ AR2 , P#0.0 ];

         L     #Mem_Accu2;
         L     #Mem_Accu1;
         LAR1  #Mem_AR1;  // Recuperar AR1
         LAR2  #Mem_AR2;  // Recuperar AR2
   next: NOP   0;
   // Fin

         JU    Bucle_1;

   Bucle_2:L     #Length_Filas_CapaReceta_DB;
         SLD   3;
         +AR1;
         L     #Length_Filas_CapaReceta_DI;
         SLD   3;
         +AR2;
         L     0;

   Bucle_1:+AR1;
         +AR2;

         OPN   "DB_RECETAS";
         OPNDI "DB_Receta_Actual";

         AN    #Reset_Bit;
         A     DBX [ AR1 , P#0.0 ];
         =     DIX [ AR2 , P#0.0 ];

         AN    #Reset_Bit;
         A     DBX [ AR1 , P#2.0 ];
         =     DIX [ AR2 , P#2.0 ];

         A     #Primer_Elemento;
         =     DIX [ AR2 , P#4.0 ];
         R     #Primer_Elemento;


         L     #Contador_Elementos;
         L     1;
         +I;
         T     #Contador_Elementos;
         L     #Max_Nro_Elementos;
         <I;
         L     1;
         JC    Bucle_1;

   //Apunta al elemento 1
         L     #Max_Nro_Elementos;
         L     1;
         -I;
         NEGI;
         +AR1;
         +AR2;
         L     0;
         T     #Contador_Elementos;

         L     #Contador_Filas;
         L     1;
         +I;
         T     #Contador_Filas;
         L     #Max_Nro_Filas;
         <I;
         JC    Bucle_2;

   //Determinar qué capa se debe cargar a continuación
         L     #"Nro CapaActual";
         INC   1;
         T     #"Nro CapaActual";
         L     #Max_Nro_Capas;
         <I;
         JC    Ok_1;
         L     1;
         T     "Proceso Dosificador".Capa_Actual;


         L     1;
         T     "Proceso Dosificador".Capa_Actual;
         T     "Proceso Empujador".Capa_Actual;



         BEU;  // Acá sale del bloque


   Ok_1: NOP   0;  // No se terminaron las capas
         L     #"Nro CapaActual";
         L     #Nro_Capas;
         <I;
         JC    Ok_2;
   // BEA
         L     #Índice_Capa_DI;
         L     1;
         +I;
         T     #Índice_Capa_DI;
         SET;
         S     #Reset_Bit;
         JU    Bucle_3;
   Ok_2: NOP   0;  // No se terminaron las capas válidas
         L     #"Nro CapaActual";
         L     #Nro_CapasDistintas;
         MOD;
         T     #índice_Capa_DB;
         L     #Índice_Capa_DI;
         L     1;
         +I;
         T     #Índice_Capa_DI;
         JU    Bucle_3;

   m000: NOP   0;
END_REGION

REGION Network 8: Transferir Velocidad Cinta Verde de la receta
         L     #Adress_Receta;
         L     #Offset_Vel_Dosificador;
         +I;
         SLD   3;
         LAR1;
         OPN   "DB_RECETAS";
         L     DBD [ AR1 , P#0.0];
         T     "DB_Velocidades".Dosif_Vel_Ráp;
END_REGION
END_FUNCTION

FUNCTION "CAPA Proceso_Animación" : Void   // FC18, STL
{ S7_Optimized_Access := 'FALSE' }
VERSION : 0.1
BEGIN

REGION Network 1: Constantes
         L     "Proceso Empujador".Capa_Actual;
         T     #Capa_Actual;
         L     38;
         T     #Length_Capas;
         L     54;
         T     #Offset_Capas;
         L     6;
         T     #Length_Filas_DB;
         L     0;
         T     #Offset_Filas_DB;
         L     1;
         T     #Length_Elementos_DB_bit;
         L     0;
         T     #Offset_Elementos_DB_bit;

         L     1;
         T     #Índice_Filas;
         T     #Índice_Elementos;

         SET;
         R     #f_Selec;

         L     "Puntero".Length_Filas_HMI;
         T     #Length_Filas_DI;
         L     "Puntero".Offset_Filas_HMI;
         T     #Offset_Filas_DI;
         L     "Puntero".Length_Elementos_HMI;
         T     #Length_Elementos_DI;
         L     "Puntero".Offset_Elementos_HMI;
         T     #Offset_Elementos_DI;

         L     "Constante".Elemento_PRESENTE;
         T     #Elemento_Cargado;
         L     "Constante".Elemento_SELECCIONADO;
         T     #Elemento_Siguiente;
         L     "Constante".Elemento_AUSENTE;
         T     #Elemento_Ausente;

         L     "Puntero".Max_Nro_Elementos;
         T     #Max_Nro_Elementos;
         L     "Puntero".Max_Nro_Filas;
         T     #Max_Nro_Filas;
END_REGION

